// TIA Portal project "EbAndon v3_0_16" (V15) (continued)

VAR_GLOBAL   // PLC tag table "BFL 03"
   "BFL 03 IO" AT %QD1080 : DWord;
   "BFL 03 KP8 In" AT %ID80 : DWord;
   "BFL 03 KP8 Out" AT %QD80 : DWord;
END_VAR

VAR_GLOBAL   // PLC tag table "LGS 01"
   "LGS 01 IO" AT %QD1084 : DWord;
   "LGS 01 KP8 In" AT %ID84 : DWord;
   "LGS 01 KP8 Out" AT %QD84 : DWord;
END_VAR

VAR_GLOBAL   // PLC tag table "LGS 02"
   "LGS 02 IO" AT %QD1088 : DWord;
   "LGS 02 KP8 In" AT %ID88 : DWord;
   "LGS 02 KP8 Out" AT %QD88 : DWord;
END_VAR

VAR_GLOBAL   // PLC tag table "CHM 01"
   "CHM 01 IO" AT %QD1092 : DWord;
   "CHM 01 KP8 In" AT %ID92 : DWord;
   "CHM 01 KP8 Out" AT %QD92 : DWord;
END_VAR

VAR_GLOBAL CONSTANT   // PLC tag table "Comm Diag"
   "pnioDeviceCount" : Int := 48;   // Upper limit of devices per HMI screen
   "USERDIAG_SLOTS_PER_SCREEN_UPPER_LIM" : Int := 31;   // Upper limit of slots per HMI screen
   "USERDIAG_SLOTS_PER_DEVICE_UPPER_LIM" : Int := 31;   // max number of modules per device
   "USERDIAG_DEVICES_PER_IO_SYSTEM_UPPER_LIM" : Int := 128;   // Upper limit of devices/slaves per IO-System/DP-Mastersystem
   "USERDIAG_SLOTS_PER_PLC_UPPER_LIM" : Int := 31;   // max number of local modules
   "USERDIAG_IO_SYSTEMS_UPPER_LIM" : Int := 1;   // Upper limit of IO-Systems/DP-Mastersystems
   "USERDIAG_IOSYSTEM_1" : Int := 1;   // Index for first IO-System/DP-Mastersystem
END_VAR

VAR_GLOBAL CONSTANT   // PLC tag table "Color Library"
   "BkBk" : USInt := 0;
   "BgWh" : USInt := 1;
   "FgWh" : USInt := 2;
   "FlWh" : USInt := 3;
   "BgGray" : USInt := 4;
   "FgGray" : USInt := 5;
   "FlGray" : USInt := 6;
   "BgLRd" : USInt := 7;
   "FgLRd" : USInt := 8;
   "FlLRd" : USInt := 9;
   "BgDRd" : USInt := 10;
   "FgDRd" : USInt := 11;
   "FlDrd" : USInt := 12;
   "BgLYe" : USInt := 13;
   "FgLYe" : USInt := 14;
   "FlLYe" : USInt := 15;
   "BgDYe" : USInt := 16;
   "FgDYe" : USInt := 17;
   "FlDYe" : USInt := 18;
   "BgLGr" : USInt := 19;
   "FgLGr" : USInt := 20;
   "FlLGr" : USInt := 21;
   "BgDGr" : USInt := 22;
   "FgDGr" : USInt := 23;
   "FlDGr" : USInt := 24;
   "BgLTe" : USInt := 25;
   "FgLTe" : USInt := 26;
   "FlLTe" : USInt := 27;
   "BgDTe" : USInt := 28;
   "FgDTe" : USInt := 29;
   "FlDTe" : USInt := 30;
   "BgLBl" : USInt := 31;
   "FgLBl" : USInt := 32;
   "FlLBl" : USInt := 33;
   "BgDBl" : USInt := 34;
   "FgDBl" : USInt := 35;
   "FlDBl" : USInt := 36;
   "BgLPu" : USInt := 37;
   "FgLPu" : USInt := 38;   // foreground light purple
   "FlLPu" : USInt := 39;
   "BgDPu" : USInt := 40;
   "FgDPu" : USInt := 41;
   "FlDPu" : USInt := 42;
   "disabled" : USInt := 254;
   "invisible" : USInt := 255;
   "LBlDRd" : USInt := 43;
   "DRdLBl" : USInt := 44;
   "LBlDRdFl" : USInt := 45;
   "DBlDRd" : USInt := 46;
   "DRdDBl" : USInt := 47;
   "DBlDRdFl" : USInt := 48;
END_VAR

VAR_GLOBAL CONSTANT   // PLC tag table "Station Meta Data"
   "ptsPerStn" : Int := 7;
   "stnCount" : Int := 30;
   "defaultAlotted" : Real := 1800.0;
   "defaultCritical" : Real := 300.0;
   "menuCntPerStn" : Int := 49;
   "mStringLen" : Int := 40;
   "sStringLen" : Int := 20;
   "lStringLen" : Int := 60;
END_VAR

VAR_GLOBAL   // PLC tag table "Simulation"
   "simMode" AT %M100.3 : Bool;
END_VAR

VAR_GLOBAL CONSTANT   // PLC tag table "Simulation"
   "simKP8Count" : Int := 11;
END_VAR

VAR_GLOBAL CONSTANT   // PLC tag table "Station IDs"
   "VOLVO 16 01" : Int := 0;
   "VOLVO 16 02" : Int := 1;
   "VOLVO 16 03" : Int := 2;
   "VOLVO 16 04" : Int := 3;
   "VOLVO 16 05" : Int := 4;
   "VOLVO 16 06" : Int := 5;
   "VOLVO 16 07" : Int := 6;
   "VOLVO 16 08" : Int := 7;
   "VOLVO 16 09" : Int := 8;
   "VOLVO 16 10" : Int := 9;
   "VOLVO 16 11" : Int := 10;
   "CHM 01" : Int := 11;
   "CHM 02" : Int := 12;
   "CHM 03" : Int := 13;
   "CHM 04" : Int := 14;
   "CHM 05" : Int := 15;
   "CDO 01" : Int := 16;
   "CDO 02" : Int := 17;
   "CDO 03" : Int := 18;
   "BFL 01" : Int := 19;
   "BFL 02" : Int := 20;
   "BFL 03" : Int := 21;
   "LGS 01" : Int := 22;
   "LGS 02" : Int := 23;
   "LGS 03" : Int := 24;
   "CV 01" : Int := 25;
   "CV 02" : Int := 26;
   "CV 03" : Int := 27;
   "CV 04" : Int := 28;
   "PC 01" : Int := 29;
   "PC 02" : Int := 30;
END_VAR

VAR_GLOBAL CONSTANT   // PLC tag table "LED Sign"
   "ledRowCount" : Int := 11;
END_VAR

VAR_GLOBAL CONSTANT   // PLC tag table "HMI Part Request Screen"
   "partReqHmiRowCount" : Int := 11;   // number of rows displayed on hmi
END_VAR

VAR_GLOBAL CONSTANT   // PLC tag table "HMI Settings Screen"
   "hmiSelStnCount" : Int := 11;   // labels for settings screen
END_VAR

VAR_GLOBAL CONSTANT   // PLC tag table "Part Request Data Base"
   "partReqDataRowCount" : Int := 199;
END_VAR

VAR_GLOBAL CONSTANT   // PLC tag table "HMI Select Station"
   "hmiStnCount" : Int := 4;   // number of stations using basic panel instead of kp8 (-1 for array)
   "hmiStnMenuSelScrnBtnCnt" : Int := 29;   // number of buttons on menu select screen (short and long rows use different data, -1 for array)
   "hmiStnMenuSelLblCnt" : Int := 29;   // number of labels (2 per row, short & long rows use same data, - 1 for array)
   "hmiStnPartSelScrnBtnCnt" : Int := 7;   // number of buttons on part select screen (-1 for array)
   "hmiStnTmpltBtnCnt" : Int := 1;   // number of button on the template (-1 for array)
END_VAR

VAR_GLOBAL   // PLC tag table "LGS 03"
   "LGS 03 IO" AT %QD1096 : DWord;
   "LGS 03 KP8 In" AT %ID96 : DWord;
   "LGS 03 KP8 Out" AT %QD96 : DWord;
END_VAR

VAR_GLOBAL   // PLC tag table "CV 01"
   "CV 01 IO" AT %QD1100 : DWord;
   "CV 01 KP8 In" AT %ID100 : DWord;
   "CV 01 KP8 Out" AT %QD100 : DWord;
END_VAR

VAR_GLOBAL   // PLC tag table "CV 02"
   "CV 02 IO" AT %QD1104 : DWord;
   "CV 02 KP8 In" AT %ID104 : DWord;
   "CV 02 KP8 Out" AT %QD104 : DWord;
END_VAR

VAR_GLOBAL   // PLC tag table "CV 03"
   "CV 03 IO" AT %QD1108 : DWord;
   "CV 03 KP8 In" AT %ID108 : DWord;
   "CV 03 KP8 Out" AT %QD108 : DWord;
END_VAR

VAR_GLOBAL   // PLC tag table "CV 04"
   "CV 04 IO" AT %QD1112 : DWord;
   "CV 04 KP8 In" AT %ID112 : DWord;
   "CV 04 KP8 Out" AT %QD112 : DWord;
END_VAR

VAR_GLOBAL   // PLC tag table "PC 01"
   "PC 01 IO" AT %QD1116 : DWord;
   "PC 01 KP8 In" AT %ID116 : DWord;
   "PC 01 KP8 Out" AT %QD116 : DWord;
END_VAR

VAR_GLOBAL   // PLC tag table "PC 02"
   "PC 02 IO" AT %QD1120 : DWord;
   "PC 02 KP8 In" AT %ID120 : DWord;
   "PC 02 KP8 Out" AT %QD120 : DWord;
END_VAR

TYPE "Stations"
   STRUCT
      me : Array[0.."stnCount"] of "Station";
   END_STRUCT;
END_TYPE

TYPE "Part Call Screen"
   STRUCT
      row : Array[0.."partReqHmiRowCount"] of "Table Row";
   END_STRUCT;
END_TYPE

TYPE "Part Req Log Row"
   STRUCT
      address : Int;
      reqType : Int;
      timeStamp : DTL;
   END_STRUCT;
END_TYPE

TYPE "Barcode Screen"
   STRUCT
      partNumber : WString[40];
      barcode : String;
      orderCancelled : Bool;
      ordered : Bool;
   END_STRUCT;
END_TYPE

TYPE "Table Row"
   STRUCT
      address : UInt;
      ordered : Bool;
      pbSelection : Struct
         actuate : Bool;
         animate : USInt;
      END_STRUCT;
      rtBackground : Struct
         animate : USInt;
      END_STRUCT;
      tfDropZone : Struct
         animate : USInt;
         value : WString[20];
      END_STRUCT;
      tfLine : Struct
         animate : USInt;
         value : WString[20];
      END_STRUCT;
      tfPartNumber : Struct
         animateDL : USInt;
         animateSL : USInt;
         value : WString[40];
      END_STRUCT;
      tfTime : Struct
         animate : USInt;
         value : WString[20];
      END_STRUCT;
   END_STRUCT;
END_TYPE

TYPE "Runtime Data"
   STRUCT
      asReal : Real;
      elapsed : LReal;
      mem : LReal;
   END_STRUCT;
END_TYPE

TYPE "KP8 Button Config"
   STRUCT
      activate : Array[0.."ptsPerStn"] of Bool;
      colorOn1 : Array[0.."ptsPerStn"] of String[10];
      colorOn2 : Array[0.."ptsPerStn"] of String[10];
      colorOff : Array[0.."ptsPerStn"] of String[10];
      flash : Array[0.."ptsPerStn"] of Bool;
      group : Array[0.."ptsPerStn"] of Int;
      mode : Array[0.."ptsPerStn"] of Bool;
   END_STRUCT;
END_TYPE

TYPE "Elapsed Time"
   STRUCT
      partReq : Array[0.."ptsPerStn"] of Real;
      resetReq : Real;
   END_STRUCT;
END_TYPE

TYPE "Part Request Data"
   STRUCT
      row : Array[0.."partReqDataRowCount"] of "Table Row";
   END_STRUCT;
END_TYPE

TYPE "Station"
   STRUCT
      animations : Array[0.."ptsPerStn"] of Int;
      btnStates : Array[0.."ptsPerStn"] of Bool;
      dropZone : USInt;
      elapsedTime : "Elapsed Time";
      groupSelect : Int;
      kp8Config : "KP8 Button Config";
      kp8In : Byte;
      kp8Out : DWord;
      init : "Station Initialization";
      line : WString[20];
      partNumbers : Array[0.."ptsPerStn"] of WString["mStringLen"];
      partOrdered : Array[0.."ptsPerStn"] of Bool;
      partRequested : Array[0.."ptsPerStn"] of Bool;
      presetTime : "Preset Time";
      settings : "Station Settings Screen";
      stackLightOut : DWord;
   END_STRUCT;
END_TYPE

TYPE "Settings"
   STRUCT
      alotted : Struct
         assign : "PB Data: Text Label";
         ioField : "IO Field Data: Timers";
      END_STRUCT;
      critical : Struct
         assign : "PB Data: Text Label";
         ioField : "IO Field Data: Timers";
      END_STRUCT;
      kp8 : Struct
         selectButtons : "PB Data: Text Label";
         btnSelState : Array[0.."ptsPerStn"] of Bool;
         buttons : Array[0.."ptsPerStn"] of "PB Data: Text Label";
         selBtnNumber : Int;
         selCount : Int;
      END_STRUCT;
      stations : Struct
         selectAll : "PB Data: Text Label";
         nextGroup : "PB Data: Graphic/Text List";
         prevGroup : "PB Data: Graphic/Text List";
         selectBtns : Array[0.."hmiSelStnCount"] of "PB Data: Text Label";
         selCount : Int;
         selNumber : Int;
      END_STRUCT;
      partNumber : Struct
         assign : "PB Data: Text Label";
         ioField : "IO Field Data: Part Number";
      END_STRUCT;
      viewingStation : Struct
         btns : Array[0.."ptsPerStn"] of "Station Assignment: Button Details";
         dzData : "Drop Zone Data";
         lineData : "Line Label Data";
         next : "PB Data: Graphic/Text List";
         previous : "PB Data: Graphic/Text List";
         "name" : WString[20];
      END_STRUCT;
   END_STRUCT;
END_TYPE

TYPE "PB Data: Graphic/Text List"
   STRUCT
      actuate : Bool;
      animate : USInt;
      listSelect : UInt;
   END_STRUCT;
END_TYPE

TYPE "LED Sign Data"
   STRUCT
      row : Array[0.."ledRowCount"] of "Table Row";
   END_STRUCT;
END_TYPE

TYPE "PB Data: Text Label"
   STRUCT
      actuate : Bool;
      animate : USInt;
      label : WString[20];
   END_STRUCT;
END_TYPE

TYPE "Station Old Presses"
   STRUCT
      me : Array[0.."stnCount", 0.."ptsPerStn"] of Bool;
   END_STRUCT;
END_TYPE

TYPE "Station Assignment: Button Details"
   STRUCT
      alloted : Struct
         animate : USInt;
         value : WString[10];
      END_STRUCT;
      critical : Struct
         animate : USInt;
         value : WString[10];
      END_STRUCT;
      label : Struct
         animate : USInt;
         value : WString[2];
      END_STRUCT;
      partNumber : Struct
         animate : USInt;
         value : WString[40];
      END_STRUCT;
      select : Struct
         actuate : Bool;
         animate : USInt;
      END_STRUCT;
   END_STRUCT;
END_TYPE

TYPE "IO Field Data: Part Number"
   STRUCT
      animate : USInt;
      inputFinished : Bool;
      value : WString[40];
   END_STRUCT;
END_TYPE

TYPE "Line Label Data"
   STRUCT
      animate : Struct
         bg : USInt;
         ioField : USInt;
      END_STRUCT;
      inputFinished : Bool;
      value : WString[10];
   END_STRUCT;
END_TYPE

TYPE "Drop Zone Data"
   STRUCT
      animate : Struct
         bg : USInt;
         ioField : USInt;
      END_STRUCT;
      inputFinished : Bool;
      value : WString[10];
   END_STRUCT;
END_TYPE

TYPE "IO Field Data: Timers"
   STRUCT
      animate : USInt;
      inputFinished : Bool;
      value : WString[5];
   END_STRUCT;
END_TYPE

TYPE "Table Nav"
   STRUCT
      top : "PB Data: Graphic/Text List";
      pageUp : "PB Data: Graphic/Text List";
      lineUp : "PB Data: Graphic/Text List";
      lineDown : "PB Data: Graphic/Text List";
      pageDown : "PB Data: Graphic/Text List";
      bottom : "PB Data: Graphic/Text List";
   END_STRUCT;
END_TYPE

TYPE "Station Sim Data"
   STRUCT
      stn : Struct
         animate : USInt;
         label : WString[20];
      END_STRUCT;
      btn : Struct
         actuate : Byte;
         animate : Array[0..7] of USInt;
         labels : Array[0..7] of WString [4];
      END_STRUCT;
   END_STRUCT;
END_TYPE

TYPE "Simulated Stations"
   STRUCT
      down : "PB Data: Graphic/Text List";
      firstStn : Int;
      me : Array[0.."simKP8Count"] of "Station Sim Data";
      up : "PB Data: Graphic/Text List";
   END_STRUCT;
END_TYPE

TYPE "Part Req Log"
   STRUCT
      me : Array[0..99] of "Part Req Log Row";
   END_STRUCT;
END_TYPE

TYPE "UserDiag_typeSlot"
   STRUCT
      hardwareId : Hw_Io := 16#0000;   // Hardware identifier of the module which is inserted in the slot
      state : USInt := 0;   // Status of the device/slave. 1:ok; 2:faulty, 3:lost connection, 4:disabled, 5:problem, 12:was faulty, 13:was lost, 14:was disabled, 15:problem gone
      exists : Bool := FALSE;   // TRUE: Modul is existing
      configured : Bool := FALSE;   // TRUE: Modul is configured
      faulty : Bool := FALSE;   // TRUE: Modul is faulty
      problem : Bool := FALSE;   // TRUE: Modul has a problem
      disabled : Bool := FALSE;   // TRUE: Modul is disabled
      error : Bool := FALSE;   // TRUE: Error in module which is inserted in the slot
   END_STRUCT;
END_TYPE

TYPE "UserDiag_typePLC"
   STRUCT
      hardwareId : Hw_Device := 16#0000;   // Hardware identifier of the PLC
      error : Bool := FALSE;   // TRUE: Error in PLC
      actualConfiguredSlots : Int := 0;   // Number of configured local slots at PLC
      slots : Array[0.."USERDIAG_SLOTS_PER_PLC_UPPER_LIM"] of "UserDiag_typeSlot";   // Information of the PLC slots; index = slotnumber; PLC always at slot 1
   END_STRUCT;
END_TYPE

TYPE "UserDiag_typeDevice"
   STRUCT
      hardwareId : Hw_Device := 16#0000;   // Hardware identifier of the device/slave
      number : UInt := 0;   // Profinet device number/Profibus address of the slave
      "name" : WString[20] := WSTRING#'';   // Name of the device/slave
      ipAddress : IP_V4;   // IP address of the device
      state : USInt := 0;   // Status of the device/slave. 1:ok; 2:faulty, 3:lost connection, 4:disabled, 5:problem, 12:was faulty, 13:was lost, 14:was disabled, 15:problem gone
      exists : Bool := FALSE;   // TRUE: Device/slave is existing
      configured : Bool := FALSE;   // TRUE: Device/slave is configured
      faulty : Bool := FALSE;   // TRUE: Device/slave is faulty
      problem : Bool := FALSE;   // TRUE: Device/slave has a problem
      disabled : Bool := FALSE;   // TRUE: Device/slave is disabled
      error : Bool := FALSE;   // TRUE: Error in device/slave
      nextDevice : Int := 0;   // device number of next device
      actualConfiguredSlots : Int := 0;   // Number of configured slots in the device/slave
      slots : Array[0.."USERDIAG_SLOTS_PER_DEVICE_UPPER_LIM"] of "UserDiag_typeSlot";   // Slot information of a device/slave
   END_STRUCT;
END_TYPE

TYPE "UserDiag_typeIOSystem"
   STRUCT
      hardwareId : Hw_IoSystem := 16#0000;   // Hardware identifier of the IO-System/DP-Mastersystem
      number : UInt := 0;   // IO-System/DP-Mastersystem number
      error : Bool := FALSE;   // TRUE: Error in IO-System/DP-Mastersystem
      firstDevice : Int := 0;   // device number (index) of first device in IO System
      lastDevice : Int := 0;   // device number (index) of last device IO System
      actualConfiguredDevices : Int := 0;   // Number of configured devices/slaves in IO-System/DP-Mastersystem
      devices : Array[1.."USERDIAG_DEVICES_PER_IO_SYSTEM_UPPER_LIM"] of "UserDiag_typeDevice";   // Device/Slave information
   END_STRUCT;
END_TYPE

TYPE "Network Health Screen"
   STRUCT
      et200spPopUp : "Station: ET200SP Comm Debug Data";
      kp8PopUp : "Station: KP8 Comm Debug Data";
      pnioDevices : Array[1.."pnioDeviceCount"] of "PB Data: Text Label";
      selectedDevice : Int;
   END_STRUCT;
   // // pnioDevices[1] : volvo1601kp8
   // // pnioDevices[2] : volvo1601et200sp
   // // pnioDevices[3] : volvo1602kp8
   // // pnioDevices[4] : volvo1602et200sp
   // // pnioDevices[5] : volvo1603kp8
   // // pnioDevices[6] : volvo1603et200sp
   // // pnioDevices[7] : volvo1604kp8
   // // pnioDevices[8] : volvo1604et200sp
   // // pnioDevices[9] : volvo1605kp8
   // // pnioDevices[10] : volvo1605et200sp
   // // pnioDevices[11] : volvo1606kp8
   // // pnioDevices[12] : volvo1606et200sp
   // // pnioDevices[13] : volvo1607kp8
   // // pnioDevices[14] : volvo1607et200sp
   // // pnioDevices[15] : volvo1608kp8
   // // pnioDevices[16] : volvo1608et200sp
   // // pnioDevices[17] : volvo1609kp8
   // // pnioDevices[18] : volvo1609et200sp
   // // pnioDevices[19] : volvo1610kp8
   // // pnioDevices[20] : volvo1610et200sp
   // // pnioDevices[21] : volvo1611kp8
   // // pnioDevices[22] : volvo1611et200sp
   // // pnioDevices[23] : chm01kp8
   // // pnioDevices[24] : chm01et200sp
   // // pnioDevices[25] : chm02kp8
   // // pnioDevices[26] : chm02et200sp
   // // pnioDevices[27] : chm03kp8
   // // pnioDevices[28] : chm03et200sp
   // // pnioDevices[29] : chm04kp8
   // // pnioDevices[30] : chm04et200sp
   // // pnioDevices[31] : chm05kp8
   // // pnioDevices[32] : chm05et200sp
   // // pnioDevices[33] : cd001kp8
   // // pnioDevices[34] : cd001et200sp
   // // pnioDevices[35] : cd002kp8
   // // pnioDevices[36] : cd002et200sp
   // // pnioDevices[37] : cd003kp8
   // // pnioDevices[38] : cd003et200sp
   // // pnioDevices[39] : bfl01kp8
   // // pnioDevices[40] : bfl01et200sp
   // // pnioDevices[41] : bfl02kp8
   // // pnioDevices[42] : bfl02et200sp
   // // pnioDevices[43] : bfl03kp8
   // // pnioDevices[44] : bfl03et200sp
   // // pnioDevices[45] : lgs01kp8
   // // pnioDevices[46] : lgs01et200sp
   // // pnioDevices[47] : lgs02kp8
   // // pnioDevices[48] : lgs02et200sp
END_TYPE

TYPE "UserDiag_typeActIOSystem"
   STRUCT
      actIOSystemNumber : Int := 1;   // Number of actual selected IO-system/DP-Mastersystem
      actIODeviceNumbers : Array[1.."pnioDeviceCount"] of UInt;   // Device numbers/profibus addresses of actual selected IO-System/DP-Mastersystem
      actIODeviceState : Array[1.."pnioDeviceCount"] of USInt;   // State of devices/slaves in actual selected IO-System/DP-Mastersystem
      actDeviceSlotsUsed : Array[0.."USERDIAG_SLOTS_PER_SCREEN_UPPER_LIM"] of Bool;   // Used slots of actual selected device/slave
      actDeviceSlotsState : Array[0.."USERDIAG_SLOTS_PER_SCREEN_UPPER_LIM"] of USInt;   // States of actual selected device/slave
   END_STRUCT;
END_TYPE

TYPE "Station: ET200SP Comm Debug Data"
   STRUCT
      dismissPB : Bool;
      IM : "ET200SP: IM Data";
      DQ01 : "ET200SP: DQ Data";
      DQ02 : "ET200SP: DQ Data";
      DQ03 : "ET200SP: DQ Data";
      profinetName : Struct
         animate : USInt;
         label : WString[20];
      END_STRUCT;
      serverModule : "ET200SP: Server Module Data";
   END_STRUCT;
END_TYPE

TYPE "ET200SP: IM Data"
   STRUCT
      bg : USInt;
      error : USInt;
      lnk01 : USInt;
      lnk02 : USInt;
      maint : USInt;
      pwr : USInt;
      run : USInt;
   END_STRUCT;
END_TYPE

TYPE "ET200SP: DQ Data"
   STRUCT
      bg : USInt;
      bgTem : USInt;
      diag : USInt;
      pwr : USInt;
      x0 : USInt;
      x1 : USInt;
      x2 : USInt;
      x3 : USInt;
      x4 : USInt;
      x5 : USInt;
      x6 : USInt;
      x7 : USInt;
   END_STRUCT;
END_TYPE

TYPE "ET200SP: Server Module Data"
   STRUCT
      bg : USInt;
   END_STRUCT;
END_TYPE

TYPE "Station: KP8 Comm Debug Data"
   STRUCT
      dismissPB : Bool;
      profinetName : Struct
         animate : USInt;
         label : WString[20];
      END_STRUCT;
      stencilBackground : USInt;
      X1P1 : Struct
         transmit : USInt;
         receive : USInt;
      END_STRUCT;
      X1P2 : Struct
         transmit : USInt;
         receive : USInt;
      END_STRUCT;
   END_STRUCT;
END_TYPE

TYPE "Station Initialization"
   STRUCT
      hard : Bool;
      soft : Bool;
   END_STRUCT;
END_TYPE

TYPE "Preset Time"
   STRUCT
      allotted : Array[0.."ptsPerStn"] of Real;
      critical : Array[0.."ptsPerStn"] of Real;
   END_STRUCT;
END_TYPE

TYPE "Station Settings Screen"
   STRUCT
      selected : Bool;
      btnSelection : Array[0.."ptsPerStn"] of Bool;
   END_STRUCT;
END_TYPE

// folder: HMI Selection Station

TYPE "HSS: Part Selection Screen"
   STRUCT
      animate : Array[0.."hmiStnPartSelScrnBtnCnt"] of Int;
      pbs : DWord;
      txt : Array[0.."hmiStnPartSelScrnBtnCnt"] of WString [40];
   END_STRUCT;
END_TYPE

TYPE "HSS: Compressed"
   STRUCT
      scrnSlctPrt : "HSS: Part Selection Screen";
      scrnSlctMn : "HSS: Menu Selection Screen";
      scrnTmplt : "HSS: Template Screen";
   END_STRUCT;
END_TYPE

TYPE "HSS: Menu Selection Screen"
   STRUCT
      animate : Array[0.."hmiStnMenuSelScrnBtnCnt"] of Int;
      pbs : DWord;
      txt : Array[0.."hmiStnMenuSelLblCnt"] of WString ["lStringLen"];
   END_STRUCT;
END_TYPE

TYPE "HSS: Template Screen"
   STRUCT
      animate : Array[0.."hmiStnTmpltBtnCnt"] of Int;
      pb : DWord;
      text : Array[0.."hmiStnTmpltBtnCnt"] of WString ["lStringLen"];
   END_STRUCT;
END_TYPE

// folder: Recipe System

TYPE "Recipe: Libraries"
   STRUCT
      stations : Array[0.."stnCount"] of "Recipe: Library";
   END_STRUCT;
END_TYPE

TYPE "Recipe: Library"
   STRUCT
      size : Int;
      wip : Array[0.."menuCntPerStn"] of WString["lStringLen"];
      raw : Array[0.."menuCntPerStn", 0.."ptsPerStn"] of WString["mStringLen"];
   END_STRUCT;
END_TYPE

// folder: (top level)

DATA_BLOCK "dbgRows"   // DB10
{ S7_Optimized_Access := 'TRUE' }
VERSION : 0.1
   VAR
      rows : Array[0..99] of DInt;
      scatterResult : Array[0..31] of Bool;
   END_VAR
BEGIN
END_DATA_BLOCK

// folder: Global Data

DATA_BLOCK "EMP IDB"   // DB1
{ S7_Optimized_Access := 'TRUE' }
VERSION : 0.1
// stored: InstanceOfName EMP
"EMP"
BEGIN
   stations.me[0].line := WSTRING#'VOLVO 16';
   stations.me[1].line := WSTRING#'VOLVO 16';
   stations.me[2].line := WSTRING#'VOLVO 16';
   stations.me[0].dropZone := 1;
   stations.me[1].dropZone := 2;
   stations.me[2].dropZone := 3;
   stations.me[3].dropZone := 4;
   stations.me[3].line := WSTRING#'VOLVO 16';
   stations.me[4].dropZone := 5;
   stations.me[4].line := WSTRING#'VOLVO 16';
   stations.me[5].line := WSTRING#'VOLVO 16';
   stations.me[5].dropZone := 6;
   stations.me[6].dropZone := 7;
   stations.me[6].line := WSTRING#'VOLVO 16';
   stations.me[7].dropZone := 8;
   stations.me[7].line := WSTRING#'VOLVO 16';
   stations.me[8].dropZone := 9;
   stations.me[8].line := WSTRING#'VOLVO 16';
   stations.me[9].dropZone := 10;
   stations.me[9].line := WSTRING#'VOLVO 16';
   stations.me[10].dropZone := 11;
   stations.me[10].line := WSTRING#'VOLVO 16';
   stations.me[11].line := WSTRING#'CHM';
   stations.me[11].dropZone := 1;
   stations.me[12].line := WSTRING#'CHM';
   stations.me[12].dropZone := 2;
   stations.me[13].line := WSTRING#'CHM';
   stations.me[13].dropZone := 3;
   stations.me[14].dropZone := 4;
   stations.me[14].line := WSTRING#'CHM';
   stations.me[15].line := WSTRING#'CHM';
   stations.me[15].dropZone := 5;
   stations.me[16].dropZone := 1;
   stations.me[16].line := WSTRING#'CDO';
   stations.me[17].dropZone := 2;
   stations.me[17].line := WSTRING#'CDO';
   stations.me[18].line := WSTRING#'CDO';
   stations.me[18].dropZone := 3;
   stations.me[19].dropZone := 1;
   stations.me[19].line := WSTRING#'BFL';
   stations.me[20].dropZone := 2;
   stations.me[20].line := WSTRING#'BFL';
   stations.me[21].line := WSTRING#'BFL';
   stations.me[21].dropZone := 3;
   stations.me[22].dropZone := 1;
   stations.me[22].line := WSTRING#'LGS';
   stations.me[23].line := WSTRING#'LGS';
   stations.me[23].dropZone := 2;
   stations.me[0].partNumbers[0] := WSTRING#'';
   stations.me[0].partNumbers[1] := WSTRING#'';
   stations.me[0].partNumbers[2] := WSTRING#'';
   stations.me[0].partNumbers[3] := WSTRING#'16.32.112.500.220A';
   stations.me[0].partNumbers[4] := WSTRING#'';
   stations.me[0].partNumbers[5] := WSTRING#'';
   stations.me[0].partNumbers[6] := WSTRING#'';
   stations.me[0].partNumbers[7] := WSTRING#'16.32.112.500.100A';
   stations.me[1].partNumbers[0] := WSTRING#'';
   stations.me[1].partNumbers[1] := WSTRING#'';
   stations.me[1].partNumbers[2] := WSTRING#'16.32.112.509.070A';
   stations.me[1].partNumbers[3] := WSTRING#'16.32.112.704.000C';
   stations.me[1].partNumbers[4] := WSTRING#'';
   stations.me[1].partNumbers[5] := WSTRING#'';
   stations.me[1].partNumbers[6] := WSTRING#'16.32.112.504.060A';
   stations.me[1].partNumbers[7] := WSTRING#'16.32.112.500.060D';
   stations.me[2].partNumbers[0] := WSTRING#'';
   stations.me[2].partNumbers[1] := WSTRING#'16.32.112.509.050E';
   stations.me[2].partNumbers[2] := WSTRING#'16.32.112.504.070G';
   stations.me[2].partNumbers[3] := WSTRING#'16.32.112.851.001A';
   stations.me[2].partNumbers[4] := WSTRING#'';
   stations.me[2].partNumbers[5] := WSTRING#'16.32.112.509.080F';
   stations.me[2].partNumbers[6] := WSTRING#'16.32.112.870.000C';
   stations.me[2].partNumbers[7] := WSTRING#'16.32.112.851.000A';
   stations.me[3].partNumbers[0] := WSTRING#'';
   stations.me[3].partNumbers[1] := WSTRING#'16.32.112.522.130A';
   stations.me[3].partNumbers[2] := WSTRING#'16.32.112.522.050A';
   stations.me[3].partNumbers[3] := WSTRING#'16.32.112.521.020B';
   stations.me[3].partNumbers[4] := WSTRING#'';
   stations.me[3].partNumbers[5] := WSTRING#'16.32.112.522.040D';
   stations.me[3].partNumbers[6] := WSTRING#'16.32.112.521.010B';
   stations.me[3].partNumbers[7] := WSTRING#'16.32.112.521.030A';
   stations.me[4].partNumbers[0] := WSTRING#'';
   stations.me[4].partNumbers[1] := WSTRING#'';
   stations.me[4].partNumbers[2] := WSTRING#'';
   stations.me[4].partNumbers[3] := WSTRING#'';
   stations.me[4].partNumbers[4] := WSTRING#'';
   stations.me[4].partNumbers[5] := WSTRING#'';
   stations.me[4].partNumbers[6] := WSTRING#'';
   stations.me[4].partNumbers[7] := WSTRING#'16.32.112.529.020B';
   stations.me[5].partNumbers[0] := WSTRING#'';
   stations.me[5].partNumbers[1] := WSTRING#'16.32.112.529.010A';
   stations.me[5].partNumbers[2] := WSTRING#'16.32.112.529.030A';
   stations.me[5].partNumbers[3] := WSTRING#'16.32.112.502.060B';
   stations.me[5].partNumbers[4] := WSTRING#'';
   stations.me[5].partNumbers[5] := WSTRING#'16.32.112.529.050D';
   stations.me[5].partNumbers[6] := WSTRING#'16.32.112.502.070E';
   stations.me[5].partNumbers[7] := WSTRING#'16.32.112.502.050B';
   stations.me[6].partNumbers[0] := WSTRING#'';
   stations.me[6].partNumbers[1] := WSTRING#'16.32.112.621.020A';
   stations.me[6].partNumbers[2] := WSTRING#'16.32.112.621.010A';
   stations.me[6].partNumbers[3] := WSTRING#'16.32.112.751.000D';
   stations.me[6].partNumbers[4] := WSTRING#'';
   stations.me[6].partNumbers[5] := WSTRING#'16.32.112.751.001C';
   stations.me[6].partNumbers[6] := WSTRING#'16.32.112.601.040A';
   stations.me[6].partNumbers[7] := WSTRING#'16.32.112.601.030A';
   stations.me[7].partNumbers[0] := WSTRING#'';
   stations.me[7].partNumbers[1] := WSTRING#'';
   stations.me[7].partNumbers[2] := WSTRING#'';
   stations.me[7].partNumbers[3] := WSTRING#'16.32.112.500.520B';
   stations.me[7].partNumbers[4] := WSTRING#'';
   stations.me[7].partNumbers[5] := WSTRING#'';
   stations.me[7].partNumbers[6] := WSTRING#'16.32.112.500.090B';
   stations.me[7].partNumbers[7] := WSTRING#'16.32.112.500.120A';
   stations.me[8].partNumbers[0] := WSTRING#'';
   stations.me[8].partNumbers[1] := WSTRING#'';
   stations.me[8].partNumbers[2] := WSTRING#'';
   stations.me[8].partNumbers[3] := WSTRING#'16.32.112.580.020A';
   stations.me[8].partNumbers[4] := WSTRING#'';
   stations.me[8].partNumbers[5] := WSTRING#'';
   stations.me[8].partNumbers[6] := WSTRING#'16.32.112.500.300E';
   stations.me[8].partNumbers[7] := WSTRING#'16.32.112.520.300E';
   stations.me[9].partNumbers[0] := WSTRING#'';
   stations.me[9].partNumbers[1] := WSTRING#'';
   stations.me[9].partNumbers[2] := WSTRING#'';
   stations.me[9].partNumbers[3] := WSTRING#'16.32.112.757.001A';
   stations.me[9].partNumbers[4] := WSTRING#'';
   stations.me[9].partNumbers[5] := WSTRING#'';
   stations.me[9].partNumbers[6] := WSTRING#'';
   stations.me[9].partNumbers[7] := WSTRING#'16.32.112.757.000A';
   stations.me[10].partNumbers[0] := WSTRING#'';
   stations.me[10].partNumbers[1] := WSTRING#'';
   stations.me[10].partNumbers[2] := WSTRING#'';
   stations.me[10].partNumbers[3] := WSTRING#'16.32.112.500.150B';
   stations.me[10].partNumbers[4] := WSTRING#'';
   stations.me[10].partNumbers[5] := WSTRING#'';
   stations.me[10].partNumbers[6] := WSTRING#'16.32.806.502.080A';
   stations.me[10].partNumbers[7] := WSTRING#'16.32.112.500.160A';
   stations.me[11].partNumbers[0] := WSTRING#'';
   stations.me[11].partNumbers[1] := WSTRING#'';
   stations.me[11].partNumbers[2] := WSTRING#'';
   stations.me[11].partNumbers[3] := WSTRING#'16.08.216.515.008C';
   stations.me[11].partNumbers[4] := WSTRING#'';
   stations.me[11].partNumbers[5] := WSTRING#'';
   stations.me[11].partNumbers[6] := WSTRING#'16.08.216.181.110B';
   stations.me[11].partNumbers[7] := WSTRING#'16.08.208.131.010L';
   stations.me[12].partNumbers[0] := WSTRING#'';
   stations.me[12].partNumbers[1] := WSTRING#'16.08.216.526.009A';
   stations.me[12].partNumbers[2] := WSTRING#'16.08.216.871.010C';
   stations.me[12].partNumbers[3] := WSTRING#'16.08.216.141.010C';
   stations.me[12].partNumbers[4] := WSTRING#'';
   stations.me[12].partNumbers[5] := WSTRING#'16.08.216.526.002C';
   stations.me[12].partNumbers[6] := WSTRING#'16.08.215.871.010C';
   stations.me[12].partNumbers[7] := WSTRING#'16.08.215.141.010C';
   stations.me[13].partNumbers[0] := WSTRING#'';
   stations.me[13].partNumbers[1] := WSTRING#'';
   stations.me[13].partNumbers[2] := WSTRING#'16.08.216.251.000B';
   stations.me[13].partNumbers[3] := WSTRING#'16.08.216.911.000G';
   stations.me[13].partNumbers[4] := WSTRING#'';
   stations.me[13].partNumbers[5] := WSTRING#'';
   stations.me[13].partNumbers[6] := WSTRING#'16.08.216.911.000H';
   stations.me[13].partNumbers[7] := WSTRING#'16.08.216.911.000C';
   stations.me[14].partNumbers[0] := WSTRING#'';
   stations.me[14].partNumbers[1] := WSTRING#'';
   stations.me[14].partNumbers[2] := WSTRING#'16.08.216.181.100A';
   stations.me[14].partNumbers[3] := WSTRING#'16.08.216.910.020B';
   stations.me[14].partNumbers[4] := WSTRING#'';
   stations.me[14].partNumbers[5] := WSTRING#'16.08.216.181.090A';
   stations.me[14].partNumbers[6] := WSTRING#'16.08.216.722.001A';
   stations.me[14].partNumbers[7] := WSTRING#'16.08.216.181.010B';
   stations.me[15].partNumbers[0] := WSTRING#'';
   stations.me[15].partNumbers[1] := WSTRING#'16.08.211.551.000B';
   stations.me[15].partNumbers[2] := WSTRING#'16.08.216.511.000C';
   stations.me[15].partNumbers[3] := WSTRING#'16.08.208.501.000B';
   stations.me[15].partNumbers[4] := WSTRING#'';
   stations.me[15].partNumbers[5] := WSTRING#'16.08.216.551.000B';
   stations.me[15].partNumbers[6] := WSTRING#'16.08.216.231.000B';
   stations.me[15].partNumbers[7] := WSTRING#'16.08.216.501.000C';
   stations.me[16].partNumbers[0] := WSTRING#'';
   stations.me[16].partNumbers[1] := WSTRING#'';
   stations.me[16].partNumbers[2] := WSTRING#'';
   stations.me[16].partNumbers[3] := WSTRING#'16.08.216.911.030B';
   stations.me[16].partNumbers[4] := WSTRING#'';
   stations.me[16].partNumbers[5] := WSTRING#'';
   stations.me[16].partNumbers[6] := WSTRING#'16.08.216.912.050A';
   stations.me[16].partNumbers[7] := WSTRING#'16.08.216.912.060B$L16.08.216.202.080A';
   stations.me[17].partNumbers[0] := WSTRING#'';
   stations.me[17].partNumbers[1] := WSTRING#'';
   stations.me[17].partNumbers[2] := WSTRING#'16.08.216.790.001A';
   stations.me[17].partNumbers[3] := WSTRING#'16.08.208.691.010D';
   stations.me[17].partNumbers[4] := WSTRING#'';
   stations.me[17].partNumbers[5] := WSTRING#'';
   stations.me[17].partNumbers[6] := WSTRING#'16.08.216.501.010A';
   stations.me[17].partNumbers[7] := WSTRING#'16.08.208.531.020L';
   stations.me[18].partNumbers[0] := WSTRING#'';
   stations.me[18].partNumbers[1] := WSTRING#'';
   stations.me[18].partNumbers[2] := WSTRING#'';
   stations.me[18].partNumbers[3] := WSTRING#'16.08.216.911.040B$L16.08.216.200.050A';
   stations.me[18].partNumbers[4] := WSTRING#'';
   stations.me[18].partNumbers[5] := WSTRING#'';
   stations.me[18].partNumbers[6] := WSTRING#'16.08.216181.020A$L16.08.208.331.000F';
   stations.me[18].partNumbers[7] := WSTRING#'16.08.216.951.010A';
   stations.me[19].partNumbers[0] := WSTRING#'';
   stations.me[19].partNumbers[1] := WSTRING#'16.08.216.521.000C';
   stations.me[19].partNumbers[2] := WSTRING#'16.08.216.831.020A';
   stations.me[19].partNumbers[3] := WSTRING#'16.08.208.151.010F';
   stations.me[19].partNumbers[4] := WSTRING#'';
   stations.me[19].partNumbers[5] := WSTRING#'16.08.217.411.080A';
   stations.me[19].partNumbers[6] := WSTRING#'16.08.216.151.010B';
   stations.me[19].partNumbers[7] := WSTRING#'16.08.211.511.020F';
   stations.me[20].partNumbers[0] := WSTRING#'';
   stations.me[20].partNumbers[1] := WSTRING#'';
   stations.me[20].partNumbers[2] := WSTRING#'';
   stations.me[20].partNumbers[3] := WSTRING#'';
   stations.me[20].partNumbers[4] := WSTRING#'';
   stations.me[20].partNumbers[5] := WSTRING#'';
   stations.me[20].partNumbers[6] := WSTRING#'';
   stations.me[20].partNumbers[7] := WSTRING#'PEANUTS';
   stations.me[21].partNumbers[0] := WSTRING#'';
   stations.me[21].partNumbers[1] := WSTRING#'';
   stations.me[21].partNumbers[2] := WSTRING#'';
   stations.me[21].partNumbers[3] := WSTRING#'RINGS CART';
   stations.me[21].partNumbers[4] := WSTRING#'';
   stations.me[21].partNumbers[5] := WSTRING#'';
   stations.me[21].partNumbers[6] := WSTRING#'';
   stations.me[21].partNumbers[7] := WSTRING#'16.08.208.011.010G';
   stations.me[22].partNumbers[0] := WSTRING#'';
   stations.me[22].partNumbers[1] := WSTRING#'';
   stations.me[22].partNumbers[2] := WSTRING#'';
   stations.me[22].partNumbers[3] := WSTRING#'16.08.208.161.020F';
   stations.me[22].partNumbers[4] := WSTRING#'';
   stations.me[22].partNumbers[5] := WSTRING#'';
   stations.me[22].partNumbers[6] := WSTRING#'16.08.211.121.000G';
   stations.me[22].partNumbers[7] := WSTRING#'16.08.216.161.020A';
   stations.me[23].partNumbers[0] := WSTRING#'';
   stations.me[23].partNumbers[1] := WSTRING#'';
   stations.me[23].partNumbers[2] := WSTRING#'';
   stations.me[23].partNumbers[3] := WSTRING#'';
   stations.me[23].partNumbers[4] := WSTRING#'';
   stations.me[23].partNumbers[5] := WSTRING#'';
   stations.me[23].partNumbers[6] := WSTRING#'';
   stations.me[23].partNumbers[7] := WSTRING#'16.08.208.021.020C';
   stations.me[24].line := WSTRING#'LGS';
   stations.me[24].dropZone := 3;
   stations.me[25].dropZone := 1;
   stations.me[25].line := WSTRING#'CV';
   stations.me[26].dropZone := 2;
   stations.me[26].line := WSTRING#'CV';
   stations.me[27].dropZone := 3;
   stations.me[27].line := WSTRING#'CV';
   stations.me[28].dropZone := 4;
   stations.me[28].line := WSTRING#'CV';
   stations.me[29].dropZone := 1;
   stations.me[29].line := WSTRING#'PC';
   stations.me[30].line := WSTRING#'PC';
   stations.me[30].dropZone := 2;
   stations.me[30].partNumbers[7] := WSTRING#'16.08.216.011.030B';
END_DATA_BLOCK

DATA_BLOCK "HMI"   // DB2
{ S7_Optimized_Access := 'TRUE' }
VERSION : 0.1
   VAR
      barcode : "Barcode Screen";
      networkHealth : "Network Health Screen";
      partCall : "Part Call Screen";
      screenNumber : Int;
      settings : "Settings";
      simStations : "Simulated Stations";
      tableNav : "Table Nav";
   END_VAR
BEGIN
END_DATA_BLOCK

DATA_BLOCK "Parts"   // DB3
{ S7_Optimized_Access := 'TRUE' }
VERSION : 0.1
   VAR RETAIN
      pRow : Int;
      requests : "Part Request Data";
   END_VAR
BEGIN
END_DATA_BLOCK

DATA_BLOCK "LED Sign"   // DB4
{ S7_Optimized_Access := 'TRUE' }
VERSION : 0.1
   VAR
      request : "LED Sign Data";
   END_VAR
BEGIN
END_DATA_BLOCK

DATA_BLOCK "Log Buffer"   // DB5
{ S7_Optimized_Access := 'TRUE' }
VERSION : 0.1
   VAR RETAIN
      logFlag : Int;
      partReq : "Part Req Log";
   END_VAR
BEGIN
END_DATA_BLOCK

DATA_BLOCK "HMI Select Stations"   // DB6
{ S7_Optimized_Access := 'TRUE' }
VERSION : 0.1
   VAR
      me : Array[0.."hmiStnCount"] of "HSS: Compressed";
   END_VAR
BEGIN
END_DATA_BLOCK

